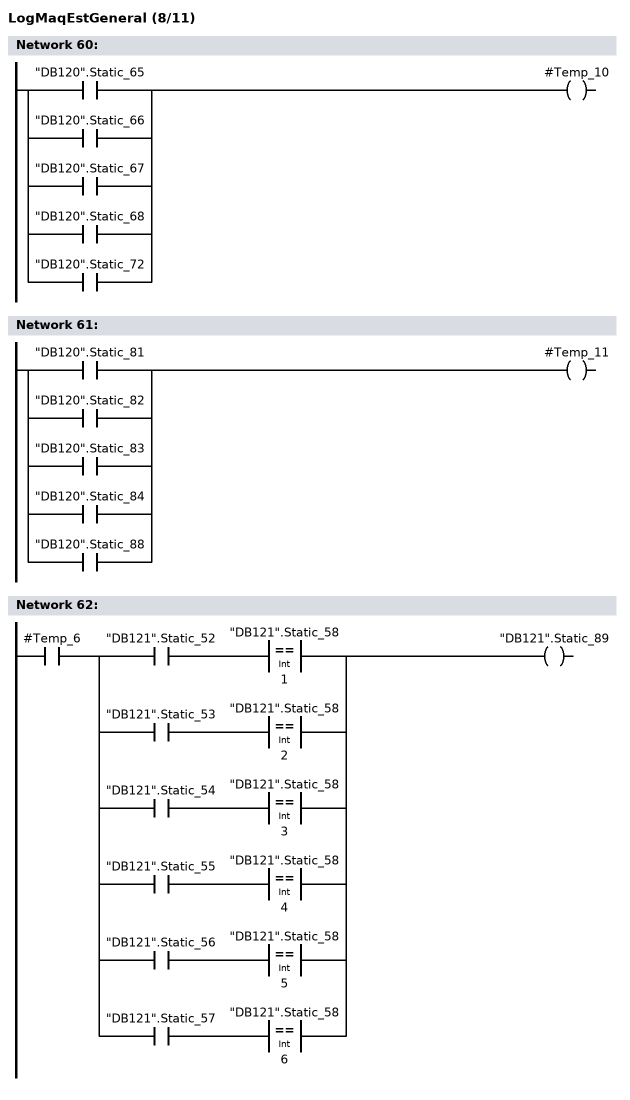
   RUNG wire#powerrail
      Contact( "DB120".Static_65 )
      wire#w1
      Coil( #Temp_10 )
   END_RUNG
   RUNG wire#powerrail
      Contact( "DB120".Static_66 )
   END_RUNG wire#w1
   RUNG wire#powerrail
      Contact( "DB120".Static_67 )
   END_RUNG wire#w1
   RUNG wire#powerrail
      Contact( "DB120".Static_68 )
   END_RUNG wire#w1
   RUNG wire#powerrail
      Contact( "DB120".Static_72 )
   END_RUNG wire#w1
   // the same network as SCL:
   #Temp_10 := "DB120".Static_65 OR "DB120".Static_66 OR "DB120".Static_67 OR "DB120".Static_68 OR "DB120".Static_72;
END_REGION

REGION Network 61
   RUNG wire#powerrail
      Contact( "DB120".Static_81 )
      wire#w1
      Coil( #Temp_11 )
   END_RUNG
   RUNG wire#powerrail
      Contact( "DB120".Static_82 )
   END_RUNG wire#w1
   RUNG wire#powerrail
      Contact( "DB120".Static_83 )
   END_RUNG wire#w1
   RUNG wire#powerrail
      Contact( "DB120".Static_84 )
   END_RUNG wire#w1
   RUNG wire#powerrail
      Contact( "DB120".Static_88 )
   END_RUNG wire#w1
   // the same network as SCL:
   #Temp_11 := "DB120".Static_81 OR "DB120".Static_82 OR "DB120".Static_83 OR "DB120".Static_84 OR "DB120".Static_88;
END_REGION

REGION Network 62
   "DB121".Static_89 := #Temp_6 AND (("DB121".Static_52 AND ("DB121".Static_58 = 1)) OR ("DB121".Static_53 AND ("DB121".Static_58 = 2)) OR ("DB121".Static_54 AND ("DB121".Static_58 = 3)) OR ("DB121".Static_55 AND ("DB121".Static_58 = 4)) OR ("DB121".Static_56 AND ("DB121".Static_58 = 5)) OR ("DB121".Static_57 AND ("DB121".Static_58 = 6)));
END_REGION

REGION Network 63
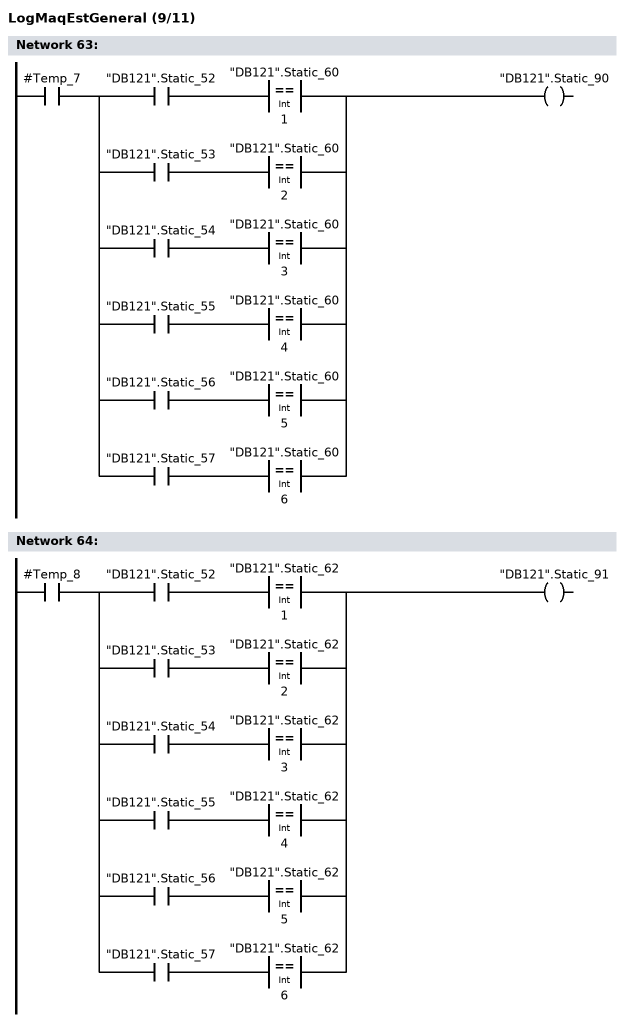
   "DB121".Static_90 := #Temp_7 AND (("DB121".Static_52 AND ("DB121".Static_60 = 1)) OR ("DB121".Static_53 AND ("DB121".Static_60 = 2)) OR ("DB121".Static_54 AND ("DB121".Static_60 = 3)) OR ("DB121".Static_55 AND ("DB121".Static_60 = 4)) OR ("DB121".Static_56 AND ("DB121".Static_60 = 5)) OR ("DB121".Static_57 AND ("DB121".Static_60 = 6)));
END_REGION

REGION Network 64
   "DB121".Static_91 := #Temp_8 AND (("DB121".Static_52 AND ("DB121".Static_62 = 1)) OR ("DB121".Static_53 AND ("DB121".Static_62 = 2)) OR ("DB121".Static_54 AND ("DB121".Static_62 = 3)) OR ("DB121".Static_55 AND ("DB121".Static_62 = 4)) OR ("DB121".Static_56 AND ("DB121".Static_62 = 5)) OR ("DB121".Static_57 AND ("DB121".Static_62 = 6)));
END_REGION

REGION Network 65
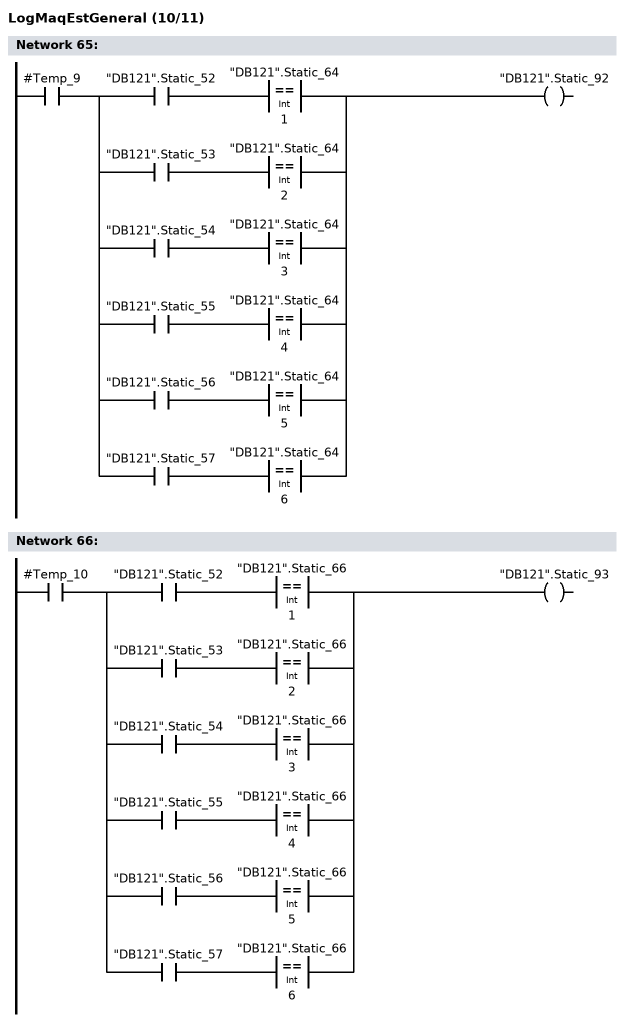
   "DB121".Static_92 := #Temp_9 AND (("DB121".Static_52 AND ("DB121".Static_64 = 1)) OR ("DB121".Static_53 AND ("DB121".Static_64 = 2)) OR ("DB121".Static_54 AND ("DB121".Static_64 = 3)) OR ("DB121".Static_55 AND ("DB121".Static_64 = 4)) OR ("DB121".Static_56 AND ("DB121".Static_64 = 5)) OR ("DB121".Static_57 AND ("DB121".Static_64 = 6)));
END_REGION

REGION Network 66
   "DB121".Static_93 := #Temp_10 AND (("DB121".Static_52 AND ("DB121".Static_66 = 1)) OR ("DB121".Static_53 AND ("DB121".Static_66 = 2)) OR ("DB121".Static_54 AND ("DB121".Static_66 = 3)) OR ("DB121".Static_55 AND ("DB121".Static_66 = 4)) OR ("DB121".Static_56 AND ("DB121".Static_66 = 5)) OR ("DB121".Static_57 AND ("DB121".Static_66 = 6)));
END_REGION

REGION Network 67
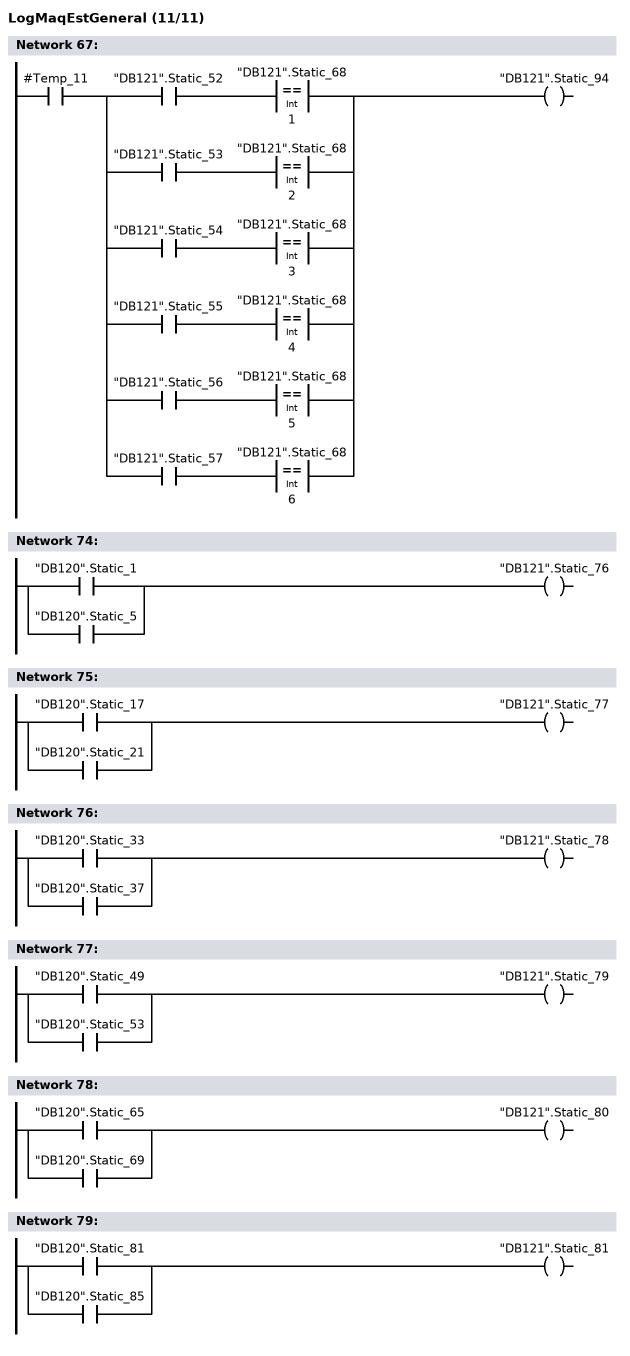
   "DB121".Static_94 := #Temp_11 AND (("DB121".Static_52 AND ("DB121".Static_68 = 1)) OR ("DB121".Static_53 AND ("DB121".Static_68 = 2)) OR ("DB121".Static_54 AND ("DB121".Static_68 = 3)) OR ("DB121".Static_55 AND ("DB121".Static_68 = 4)) OR ("DB121".Static_56 AND ("DB121".Static_68 = 5)) OR ("DB121".Static_57 AND ("DB121".Static_68 = 6)));
END_REGION

REGION Network 68 (STL)
         A(;
         L     "DB125".Static_1;
         L     1;
         ==R;
         );
         AN    "DB88".Static_12;
         O;
         A(;
         L     "DB125".Static_2;
         L     1;
         ==R;
         );
         AN    "DB88".Static_13;
         O;
         A(;
         L     "DB125".Static_3;
         L     1;
         ==R;
         );
         AN    "DB88".Static_14;
         O;
         A(;
         L     "DB125".Static_4;
         L     1;
         ==R;
         );
         AN    "DB88".Static_15;
         O;
         A(;
         L     "DB125".Static_5;
         L     1;
         ==R;
         );
         AN    "DB88".Static_16;
         O;
         A(;
         L     "DB125".Static_6;
         L     1;
         ==R;
         );
         AN    "DB88".Static_17;
         =     "DB121".Static_82;
END_REGION

REGION Network 69 (STL)
         A(;
         L     "DB125".Static_1;
         L     2;
         ==R;
         );
         AN    "DB88".Static_12;
         O;
         A(;
         L     "DB125".Static_2;
         L     2;
         ==R;
         );
         AN    "DB88".Static_13;
         O;
         A(;
         L     "DB125".Static_3;
         L     2;
         ==R;
         );
         AN    "DB88".Static_14;
         O;
         A(;
         L     "DB125".Static_4;
         L     2;
         ==R;
         );
         AN    "DB88".Static_15;
         O;
         A(;
         L     "DB125".Static_5;
         L     2;
         ==R;
         );
         AN    "DB88".Static_16;
         A(;
         L     "DB125".Static_6;
         L     2;
         ==R;
         );
         AN    "DB88".Static_17;
         =     "DB121".Static_83;
END_REGION

REGION Network 70 (STL)
         A(;
         L     "DB125".Static_1;
         L     3;
         ==R;
         );
         AN    "DB88".Static_12;
         O;
         A(;
         L     "DB125".Static_2;
         L     3;
         ==R;
         );
         AN    "DB88".Static_13;
         O;
         A(;
         L     "DB125".Static_3;
         L     3;
         ==R;
         );
         AN    "DB88".Static_14;
         O;
         A(;
         L     "DB125".Static_4;
         L     3;
         ==R;
         );
         AN    "DB88".Static_15;
         O;
         A(;
         L     "DB125".Static_5;
         L     3;
         ==R;
         );
         AN    "DB88".Static_16;
         O;
         A(;
         L     "DB125".Static_6;
         L     3;
         ==R;
         );
         AN    "DB88".Static_17;
         =     "DB121".Static_84;
END_REGION

REGION Network 71 (STL)
         A(;
         L     "DB125".Static_1;
         L     4;
         ==R;
         );
         AN    "DB88".Static_12;
         O;
         A(;
         L     "DB125".Static_2;
         L     4;
         ==R;
         );
         AN    "DB88".Static_13;
         O;
         A(;
         L     "DB125".Static_3;
         L     4;
         ==R;
         );
         AN    "DB88".Static_14;
         O;
         A(;
         L     "DB125".Static_4;
         L     4;
         ==R;
         );
         AN    "DB88".Static_15;
         O;
         A(;
         L     "DB125".Static_5;
         L     4;
         ==R;
         );
         AN    "DB88".Static_16;
         O;
         A(;
         L     "DB125".Static_6;
         L     4;
         ==R;
         );
         AN    "DB88".Static_17;
         =     "DB121".Static_85;
END_REGION

REGION Network 72 (STL)
         A(;
         L     "DB125".Static_1;
         L     5;
         ==R;
         );
         AN    "DB88".Static_12;
         O;
         A(;
         L     "DB125".Static_2;
         L     5;
         ==R;
         );
         AN    "DB88".Static_13;
         O;
         A(;
         L     "DB125".Static_3;
         L     5;
         ==R;
         );
         AN    "DB88".Static_14;
         O;
         A(;
         L     "DB125".Static_4;
         L     5;
         ==R;
         );
         AN    "DB88".Static_15;
         O;
         A(;
         L     "DB125".Static_5;
         L     5;
         ==R;
         );
         AN    "DB88".Static_16;
         O;
         A(;
         L     "DB125".Static_6;
         L     5;
         ==R;
         );
         AN    "DB88".Static_17;
         =     "DB121".Static_86;
END_REGION

REGION Network 73 (STL)
         A(;
         L     "DB125".Static_1;
         L     6;
         ==R;
         );
         AN    "DB88".Static_12;
         O;
         A(;
         L     "DB125".Static_2;
         L     6;
         ==R;
         );
         AN    "DB88".Static_13;
         O;
         A(;
         L     "DB125".Static_3;
         L     6;
         ==R;
         );
         AN    "DB88".Static_14;
         O;
         A(;
         L     "DB125".Static_4;
         L     6;
         ==R;
         );
         AN    "DB88".Static_15;
         O;
         A(;
         L     "DB125".Static_5;
         L     6;
         ==R;
         );
         AN    "DB88".Static_16;
         O;
         A(;
         L     "DB125".Static_6;
         L     6;
         ==R;
         );
         AN    "DB88".Static_17;
         =     "DB121".Static_87;
END_REGION

REGION Network 74
   RUNG wire#powerrail
      Contact( "DB120".Static_1 )
      wire#w1
      Coil( "DB121".Static_76 )
   END_RUNG
   RUNG wire#powerrail
      Contact( "DB120".Static_5 )
   END_RUNG wire#w1
   // the same network as SCL:
   "DB121".Static_76 := "DB120".Static_1 OR "DB120".Static_5;
END_REGION

REGION Network 75
   RUNG wire#powerrail
      Contact( "DB120".Static_17 )
      wire#w1
      Coil( "DB121".Static_77 )
   END_RUNG
   RUNG wire#powerrail
      Contact( "DB120".Static_21 )
   END_RUNG wire#w1
   // the same network as SCL:
   "DB121".Static_77 := "DB120".Static_17 OR "DB120".Static_21;
END_REGION

REGION Network 76
   RUNG wire#powerrail
      Contact( "DB120".Static_33 )
      wire#w1
      Coil( "DB121".Static_78 )
   END_RUNG
   RUNG wire#powerrail
      Contact( "DB120".Static_37 )
   END_RUNG wire#w1
   // the same network as SCL:
   "DB121".Static_78 := "DB120".Static_33 OR "DB120".Static_37;
END_REGION

REGION Network 77
   RUNG wire#powerrail
      Contact( "DB120".Static_49 )
      wire#w1
      Coil( "DB121".Static_79 )
   END_RUNG
   RUNG wire#powerrail
      Contact( "DB120".Static_53 )
   END_RUNG wire#w1
   // the same network as SCL:
   "DB121".Static_79 := "DB120".Static_49 OR "DB120".Static_53;
END_REGION

REGION Network 78
   RUNG wire#powerrail
      Contact( "DB120".Static_65 )
      wire#w1
      Coil( "DB121".Static_80 )
   END_RUNG
   RUNG wire#powerrail
      Contact( "DB120".Static_69 )
   END_RUNG wire#w1
   // the same network as SCL:
   "DB121".Static_80 := "DB120".Static_65 OR "DB120".Static_69;
END_REGION

REGION Network 79
   RUNG wire#powerrail
      Contact( "DB120".Static_81 )
      wire#w1
      Coil( "DB121".Static_81 )
   END_RUNG
   RUNG wire#powerrail
      Contact( "DB120".Static_85 )
   END_RUNG wire#w1
   // the same network as SCL:
   "DB121".Static_81 := "DB120".Static_81 OR "DB120".Static_85;
END_REGION
END_FUNCTION

FUNCTION "CalcEst1" : Void   // FC36, LAD
{ S7_Optimized_Access := 'FALSE' }
VERSION : 0.1
   VAR_TEMP   // added for the SCL form of the ladder/FBD networks
      _w1 : Bool;
   END_VAR
BEGIN

REGION Network 1
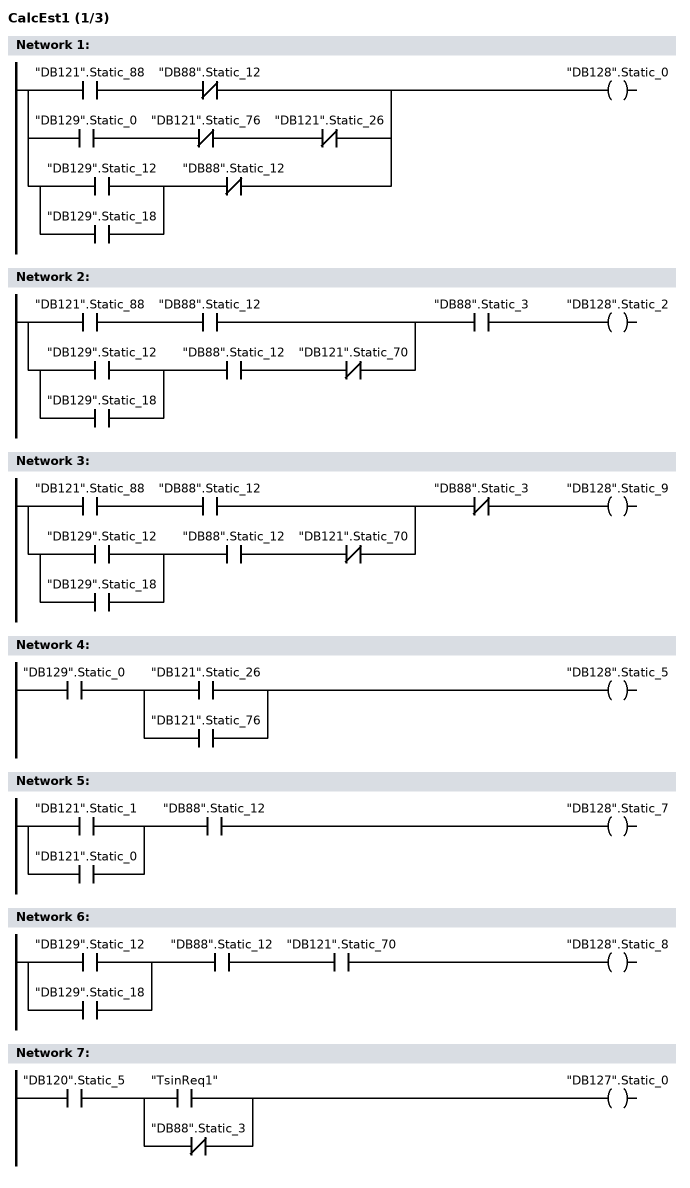
   RUNG wire#powerrail
      Contact( "DB121".Static_88 )
      I_Contact( "DB88".Static_12 )
      wire#w1
      Coil( "DB128".Static_0 )
   END_RUNG
   RUNG wire#powerrail
      Contact( "DB129".Static_0 )
      I_Contact( "DB121".Static_76 )
      I_Contact( "DB121".Static_26 )
   END_RUNG wire#w1
   RUNG wire#powerrail
      Contact( "DB129".Static_12 )
      wire#w2
      I_Contact( "DB88".Static_12 )
   END_RUNG wire#w1
   RUNG wire#powerrail
      Contact( "DB129".Static_18 )
   END_RUNG wire#w2
   // the same network as SCL:
   "DB128".Static_0 := ("DB121".Static_88 AND NOT "DB88".Static_12) OR ("DB129".Static_0 AND NOT "DB121".Static_76 AND NOT "DB121".Static_26) OR (("DB129".Static_12 OR "DB129".Static_18) AND NOT "DB88".Static_12);
END_REGION

REGION Network 2
   RUNG wire#powerrail
      Contact( "DB121".Static_88 )
      Contact( "DB88".Static_12 )
      wire#w1
      Contact( "DB88".Static_3 )
      Coil( "DB128".Static_2 )
   END_RUNG
   RUNG wire#powerrail
      Contact( "DB129".Static_12 )
      wire#w2
      Contact( "DB88".Static_12 )
      I_Contact( "DB121".Static_70 )
   END_RUNG wire#w1
   RUNG wire#powerrail
      Contact( "DB129".Static_18 )
   END_RUNG wire#w2
   // the same network as SCL:
   "DB128".Static_2 := (("DB121".Static_88 AND "DB88".Static_12) OR (("DB129".Static_12 OR "DB129".Static_18) AND "DB88".Static_12 AND NOT "DB121".Static_70)) AND "DB88".Static_3;
END_REGION

REGION Network 3
   RUNG wire#powerrail
      Contact( "DB121".Static_88 )
      Contact( "DB88".Static_12 )
      wire#w1
      I_Contact( "DB88".Static_3 )
      Coil( "DB128".Static_9 )
   END_RUNG
   RUNG wire#powerrail
      Contact( "DB129".Static_12 )
      wire#w2
      Contact( "DB88".Static_12 )
      I_Contact( "DB121".Static_70 )
   END_RUNG wire#w1
   RUNG wire#powerrail
      Contact( "DB129".Static_18 )
   END_RUNG wire#w2
   // the same network as SCL:
   "DB128".Static_9 := (("DB121".Static_88 AND "DB88".Static_12) OR (("DB129".Static_12 OR "DB129".Static_18) AND "DB88".Static_12 AND NOT "DB121".Static_70)) AND NOT "DB88".Static_3;
END_REGION

REGION Network 4
   "DB128".Static_5 := "DB129".Static_0 AND ("DB121".Static_26 OR "DB121".Static_76);
END_REGION

REGION Network 5
   RUNG wire#powerrail
      Contact( "DB121".Static_1 )
      wire#w1
      Contact( "DB88".Static_12 )
      Coil( "DB128".Static_7 )
   END_RUNG
   RUNG wire#powerrail
      Contact( "DB121".Static_0 )
   END_RUNG wire#w1
   // the same network as SCL:
   "DB128".Static_7 := ("DB121".Static_1 OR "DB121".Static_0) AND "DB88".Static_12;
END_REGION

REGION Network 6
   RUNG wire#powerrail
      Contact( "DB129".Static_12 )
      wire#w1
      Contact( "DB88".Static_12 )
      Contact( "DB121".Static_70 )
      Coil( "DB128".Static_8 )
   END_RUNG
   RUNG wire#powerrail
      Contact( "DB129".Static_18 )
   END_RUNG wire#w1
   // the same network as SCL:
   "DB128".Static_8 := ("DB129".Static_12 OR "DB129".Static_18) AND "DB88".Static_12 AND "DB121".Static_70;
END_REGION

REGION Network 7
   "DB127".Static_0 := "DB120".Static_5 AND ("TsinReq1" OR NOT "DB88".Static_3);
END_REGION

REGION Network 8
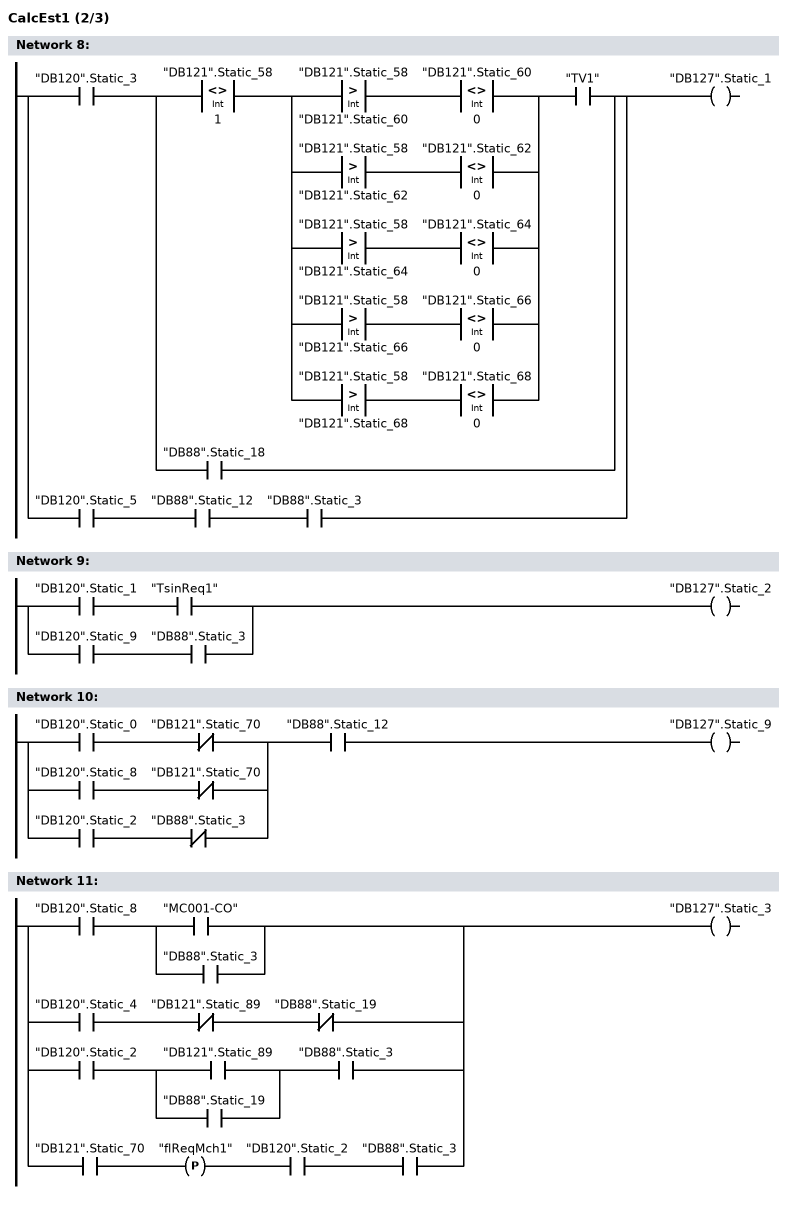
   "DB127".Static_1 := ("DB120".Static_3 AND ((("DB121".Static_58 <> 1) AND ((("DB121".Static_58 > "DB121".Static_60) AND ("DB121".Static_60 <> 0)) OR (("DB121".Static_58 > "DB121".Static_62) AND ("DB121".Static_62 <> 0)) OR (("DB121".Static_58 > "DB121".Static_64) AND ("DB121".Static_64 <> 0)) OR (("DB121".Static_58 > "DB121".Static_66) AND ("DB121".Static_66 <> 0)) OR (("DB121".Static_58 > "DB121".Static_68) AND ("DB121".Static_68 <> 0))) AND "TV1") OR "DB88".Static_18)) OR ("DB120".Static_5 AND "DB88".Static_12 AND "DB88".Static_3);
END_REGION

REGION Network 9
   RUNG wire#powerrail
      Contact( "DB120".Static_1 )
      Contact( "TsinReq1" )
      wire#w1
      Coil( "DB127".Static_2 )
   END_RUNG
   RUNG wire#powerrail
      Contact( "DB120".Static_9 )
      Contact( "DB88".Static_3 )
   END_RUNG wire#w1
   // the same network as SCL:
   "DB127".Static_2 := ("DB120".Static_1 AND "TsinReq1") OR ("DB120".Static_9 AND "DB88".Static_3);
END_REGION

REGION Network 10
   RUNG wire#powerrail
      Contact( "DB120".Static_0 )
      I_Contact( "DB121".Static_70 )
      wire#w1
      Contact( "DB88".Static_12 )
      Coil( "DB127".Static_9 )
   END_RUNG
   RUNG wire#powerrail
      Contact( "DB120".Static_8 )
      I_Contact( "DB121".Static_70 )
   END_RUNG wire#w1
   RUNG wire#powerrail
      Contact( "DB120".Static_2 )
      I_Contact( "DB88".Static_3 )
   END_RUNG wire#w1
   // the same network as SCL:
   "DB127".Static_9 := (("DB120".Static_0 AND NOT "DB121".Static_70) OR ("DB120".Static_8 AND NOT "DB121".Static_70) OR ("DB120".Static_2 AND NOT "DB88".Static_3)) AND "DB88".Static_12;
END_REGION

REGION Network 11
   #_w1 := "DB121".Static_70 AND NOT "flReqMch1";   // rising edge
   "flReqMch1" := "DB121".Static_70;
   "DB127".Static_3 := ("DB120".Static_8 AND ("MC001-CO" OR "DB88".Static_3)) OR ("DB120".Static_4 AND NOT "DB121".Static_89 AND NOT "DB88".Static_19) OR ("DB120".Static_2 AND ("DB121".Static_89 OR "DB88".Static_19) AND "DB88".Static_3) OR (#_w1 AND "DB120".Static_2 AND "DB88".Static_3);
END_REGION

REGION Network 12
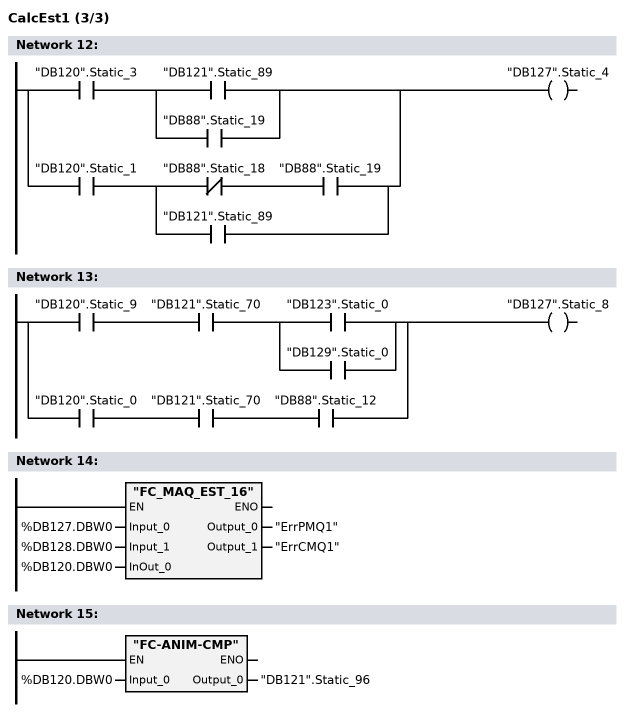
   "DB127".Static_4 := ("DB120".Static_3 AND ("DB121".Static_89 OR "DB88".Static_19)) OR ("DB120".Static_1 AND ("DB121".Static_89 OR (NOT "DB88".Static_18 AND "DB88".Static_19)));
END_REGION

REGION Network 13
   "DB127".Static_8 := ("DB120".Static_9 AND "DB121".Static_70 AND ("DB123".Static_0 OR "DB129".Static_0)) OR ("DB120".Static_0 AND "DB121".Static_70 AND "DB88".Static_12);
END_REGION

REGION Network 14
   RUNG wire#powerrail
      "FC_MAQ_EST_16"(Input_0 := %DB127.DBW0, Input_1 := %DB128.DBW0, Output_0 => "ErrPMQ1", Output_1 => "ErrCMQ1", InOut_0 := %DB120.DBW0)
   END_RUNG
   // the same network as SCL:
   "FC_MAQ_EST_16"(Input_0 := %DB127.DBW0,
                   Input_1 := %DB128.DBW0,
                   InOut_0 := %DB120.DBW0,
                   Output_0 => "ErrPMQ1",
                   Output_1 => "ErrCMQ1");
END_REGION

REGION Network 15
   RUNG wire#powerrail
      "FC-ANIM-CMP"(Input_0 := %DB120.DBW0, Output_0 => "DB121".Static_96)
   END_RUNG
   // the same network as SCL:
   "FC-ANIM-CMP"(Input_0 := %DB120.DBW0, Output_0 => "DB121".Static_96);
END_REGION
END_FUNCTION

FUNCTION "CalcEst2" : Void   // FC37, LAD
{ S7_Optimized_Access := 'FALSE' }
VERSION : 0.1
   VAR_TEMP   // added for the SCL form of the ladder/FBD networks
      _w1 : Bool;
   END_VAR
BEGIN

REGION Network 1
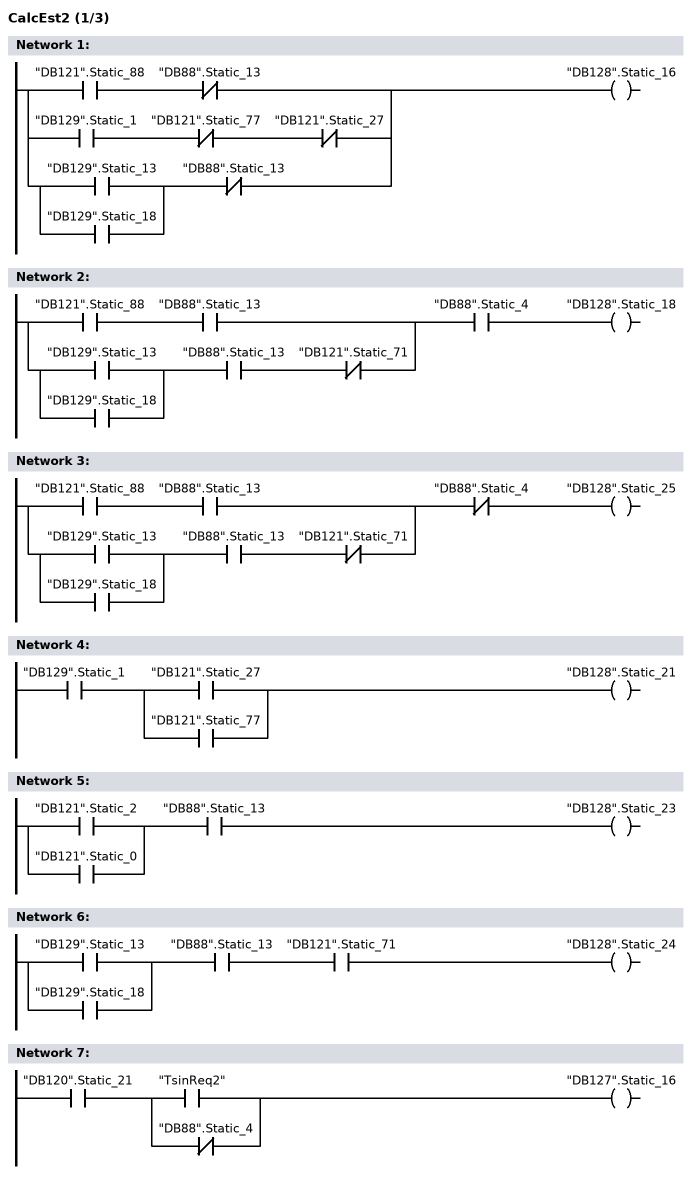
   RUNG wire#powerrail
      Contact( "DB121".Static_88 )
      I_Contact( "DB88".Static_13 )
      wire#w1
      Coil( "DB128".Static_16 )
   END_RUNG
   RUNG wire#powerrail
      Contact( "DB129".Static_1 )
      I_Contact( "DB121".Static_77 )
      I_Contact( "DB121".Static_27 )
   END_RUNG wire#w1
   RUNG wire#powerrail
      Contact( "DB129".Static_13 )
      wire#w2
      I_Contact( "DB88".Static_13 )
   END_RUNG wire#w1
   RUNG wire#powerrail
      Contact( "DB129".Static_18 )
   END_RUNG wire#w2
   // the same network as SCL:
   "DB128".Static_16 := ("DB121".Static_88 AND NOT "DB88".Static_13) OR ("DB129".Static_1 AND NOT "DB121".Static_77 AND NOT "DB121".Static_27) OR (("DB129".Static_13 OR "DB129".Static_18) AND NOT "DB88".Static_13);
END_REGION

REGION Network 2
   RUNG wire#powerrail
      Contact( "DB121".Static_88 )
      Contact( "DB88".Static_13 )
      wire#w1
      Contact( "DB88".Static_4 )
      Coil( "DB128".Static_18 )
   END_RUNG
   RUNG wire#powerrail
      Contact( "DB129".Static_13 )
      wire#w2
      Contact( "DB88".Static_13 )
      I_Contact( "DB121".Static_71 )
   END_RUNG wire#w1
   RUNG wire#powerrail
      Contact( "DB129".Static_18 )
   END_RUNG wire#w2
   // the same network as SCL:
   "DB128".Static_18 := (("DB121".Static_88 AND "DB88".Static_13) OR (("DB129".Static_13 OR "DB129".Static_18) AND "DB88".Static_13 AND NOT "DB121".Static_71)) AND "DB88".Static_4;
END_REGION

REGION Network 3
   RUNG wire#powerrail
      Contact( "DB121".Static_88 )
      Contact( "DB88".Static_13 )
      wire#w1
      I_Contact( "DB88".Static_4 )
      Coil( "DB128".Static_25 )
   END_RUNG
   RUNG wire#powerrail
      Contact( "DB129".Static_13 )
      wire#w2
      Contact( "DB88".Static_13 )
      I_Contact( "DB121".Static_71 )
   END_RUNG wire#w1
   RUNG wire#powerrail
      Contact( "DB129".Static_18 )
   END_RUNG wire#w2
   // the same network as SCL:
   "DB128".Static_25 := (("DB121".Static_88 AND "DB88".Static_13) OR (("DB129".Static_13 OR "DB129".Static_18) AND "DB88".Static_13 AND NOT "DB121".Static_71)) AND NOT "DB88".Static_4;
END_REGION

REGION Network 4
   "DB128".Static_21 := "DB129".Static_1 AND ("DB121".Static_27 OR "DB121".Static_77);
END_REGION

REGION Network 5
   RUNG wire#powerrail
      Contact( "DB121".Static_2 )
      wire#w1
      Contact( "DB88".Static_13 )
      Coil( "DB128".Static_23 )
   END_RUNG
   RUNG wire#powerrail
      Contact( "DB121".Static_0 )
   END_RUNG wire#w1
   // the same network as SCL:
   "DB128".Static_23 := ("DB121".Static_2 OR "DB121".Static_0) AND "DB88".Static_13;
END_REGION

REGION Network 6
   RUNG wire#powerrail
      Contact( "DB129".Static_13 )
      wire#w1
      Contact( "DB88".Static_13 )
      Contact( "DB121".Static_71 )
      Coil( "DB128".Static_24 )
   END_RUNG
   RUNG wire#powerrail
      Contact( "DB129".Static_18 )
   END_RUNG wire#w1
   // the same network as SCL:
   "DB128".Static_24 := ("DB129".Static_13 OR "DB129".Static_18) AND "DB88".Static_13 AND "DB121".Static_71;
END_REGION

REGION Network 7
   "DB127".Static_16 := "DB120".Static_21 AND ("TsinReq2" OR NOT "DB88".Static_4);
END_REGION

REGION Network 8
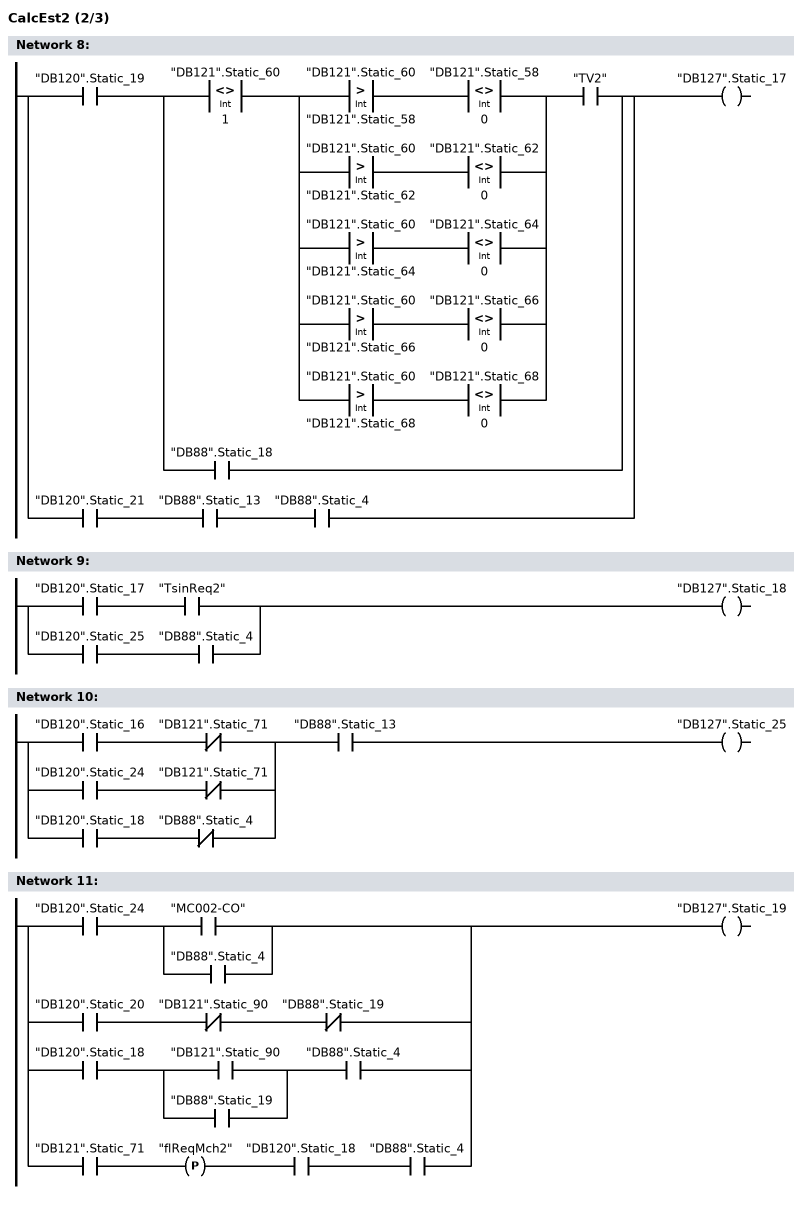
   "DB127".Static_17 := ("DB120".Static_19 AND ((("DB121".Static_60 <> 1) AND ((("DB121".Static_60 > "DB121".Static_58) AND ("DB121".Static_58 <> 0)) OR (("DB121".Static_60 > "DB121".Static_62) AND ("DB121".Static_62 <> 0)) OR (("DB121".Static_60 > "DB121".Static_64) AND ("DB121".Static_64 <> 0)) OR (("DB121".Static_60 > "DB121".Static_66) AND ("DB121".Static_66 <> 0)) OR (("DB121".Static_60 > "DB121".Static_68) AND ("DB121".Static_68 <> 0))) AND "TV2") OR "DB88".Static_18)) OR ("DB120".Static_21 AND "DB88".Static_13 AND "DB88".Static_4);
END_REGION

REGION Network 9
   RUNG wire#powerrail
      Contact( "DB120".Static_17 )
      Contact( "TsinReq2" )
      wire#w1
      Coil( "DB127".Static_18 )
   END_RUNG
   RUNG wire#powerrail
      Contact( "DB120".Static_25 )
      Contact( "DB88".Static_4 )
   END_RUNG wire#w1
   // the same network as SCL:
   "DB127".Static_18 := ("DB120".Static_17 AND "TsinReq2") OR ("DB120".Static_25 AND "DB88".Static_4);
END_REGION

REGION Network 10
   RUNG wire#powerrail
      Contact( "DB120".Static_16 )
      I_Contact( "DB121".Static_71 )
      wire#w1
      Contact( "DB88".Static_13 )
      Coil( "DB127".Static_25 )
   END_RUNG
   RUNG wire#powerrail
      Contact( "DB120".Static_24 )
      I_Contact( "DB121".Static_71 )
   END_RUNG wire#w1
   RUNG wire#powerrail
      Contact( "DB120".Static_18 )
      I_Contact( "DB88".Static_4 )
   END_RUNG wire#w1
   // the same network as SCL:
   "DB127".Static_25 := (("DB120".Static_16 AND NOT "DB121".Static_71) OR ("DB120".Static_24 AND NOT "DB121".Static_71) OR ("DB120".Static_18 AND NOT "DB88".Static_4)) AND "DB88".Static_13;
END_REGION

REGION Network 11
   #_w1 := "DB121".Static_71 AND NOT "flReqMch2";   // rising edge
   "flReqMch2" := "DB121".Static_71;
   "DB127".Static_19 := ("DB120".Static_24 AND ("MC002-CO" OR "DB88".Static_4)) OR ("DB120".Static_20 AND NOT "DB121".Static_90 AND NOT "DB88".Static_19) OR ("DB120".Static_18 AND ("DB121".Static_90 OR "DB88".Static_19) AND "DB88".Static_4) OR (#_w1 AND "DB120".Static_18 AND "DB88".Static_4);
END_REGION

REGION Network 12
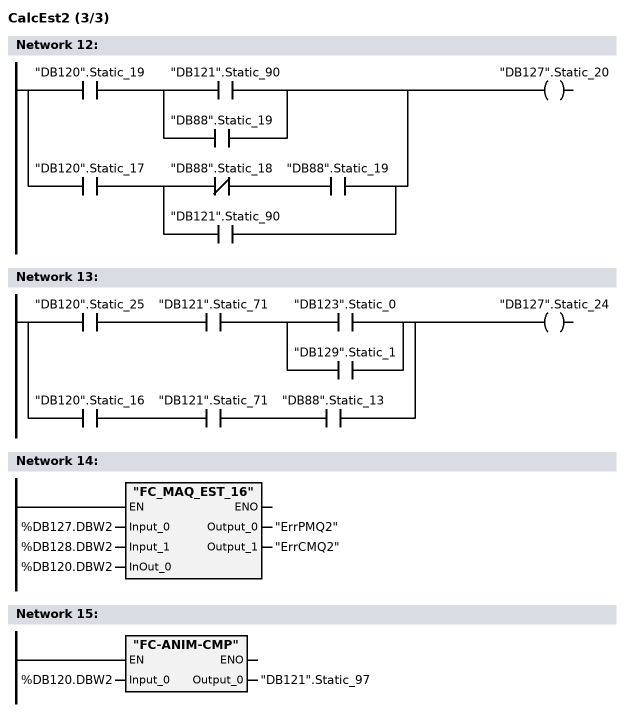
   "DB127".Static_20 := ("DB120".Static_19 AND ("DB121".Static_90 OR "DB88".Static_19)) OR ("DB120".Static_17 AND ("DB121".Static_90 OR (NOT "DB88".Static_18 AND "DB88".Static_19)));
END_REGION

REGION Network 13
   "DB127".Static_24 := ("DB120".Static_25 AND "DB121".Static_71 AND ("DB123".Static_0 OR "DB129".Static_1)) OR ("DB120".Static_16 AND "DB121".Static_71 AND "DB88".Static_13);
END_REGION

REGION Network 14
   RUNG wire#powerrail
      "FC_MAQ_EST_16"(Input_0 := %DB127.DBW2, Input_1 := %DB128.DBW2, Output_0 => "ErrPMQ2", Output_1 => "ErrCMQ2", InOut_0 := %DB120.DBW2)
   END_RUNG
   // the same network as SCL:
   "FC_MAQ_EST_16"(Input_0 := %DB127.DBW2,
                   Input_1 := %DB128.DBW2,
                   InOut_0 := %DB120.DBW2,
                   Output_0 => "ErrPMQ2",
                   Output_1 => "ErrCMQ2");
END_REGION

REGION Network 15
   RUNG wire#powerrail
      "FC-ANIM-CMP"(Input_0 := %DB120.DBW2, Output_0 => "DB121".Static_97)
   END_RUNG
   // the same network as SCL:
   "FC-ANIM-CMP"(Input_0 := %DB120.DBW2, Output_0 => "DB121".Static_97);
END_REGION
END_FUNCTION

FUNCTION "CalcEst3" : Void   // FC38, LAD
{ S7_Optimized_Access := 'FALSE' }
VERSION : 0.1
   VAR_TEMP   // added for the SCL form of the ladder/FBD networks
      _w1 : Bool;
   END_VAR
BEGIN

REGION Network 1
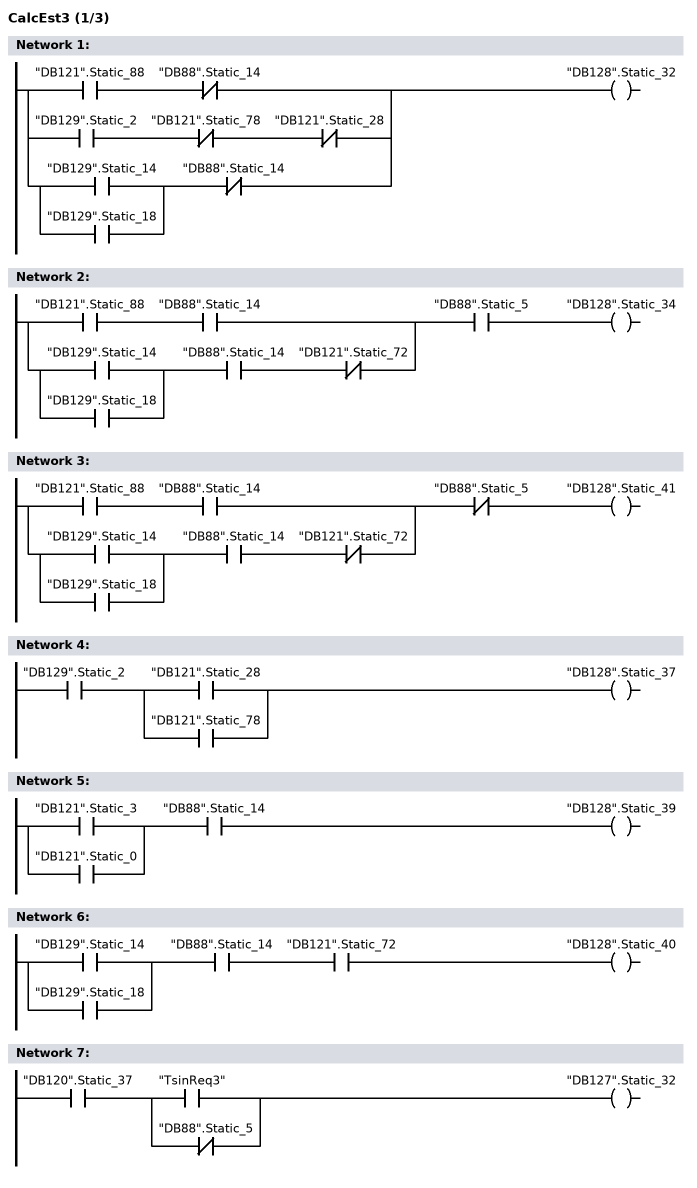
   RUNG wire#powerrail
      Contact( "DB121".Static_88 )
      I_Contact( "DB88".Static_14 )
      wire#w1
      Coil( "DB128".Static_32 )
   END_RUNG
   RUNG wire#powerrail
      Contact( "DB129".Static_2 )
      I_Contact( "DB121".Static_78 )
      I_Contact( "DB121".Static_28 )
   END_RUNG wire#w1
   RUNG wire#powerrail
      Contact( "DB129".Static_14 )
      wire#w2
      I_Contact( "DB88".Static_14 )
   END_RUNG wire#w1
   RUNG wire#powerrail
      Contact( "DB129".Static_18 )
   END_RUNG wire#w2
   // the same network as SCL:
   "DB128".Static_32 := ("DB121".Static_88 AND NOT "DB88".Static_14) OR ("DB129".Static_2 AND NOT "DB121".Static_78 AND NOT "DB121".Static_28) OR (("DB129".Static_14 OR "DB129".Static_18) AND NOT "DB88".Static_14);
END_REGION

REGION Network 2
   RUNG wire#powerrail
      Contact( "DB121".Static_88 )
      Contact( "DB88".Static_14 )
      wire#w1
      Contact( "DB88".Static_5 )
      Coil( "DB128".Static_34 )
   END_RUNG
   RUNG wire#powerrail
      Contact( "DB129".Static_14 )
      wire#w2
      Contact( "DB88".Static_14 )
      I_Contact( "DB121".Static_72 )
   END_RUNG wire#w1
   RUNG wire#powerrail
      Contact( "DB129".Static_18 )
   END_RUNG wire#w2
   // the same network as SCL:
   "DB128".Static_34 := (("DB121".Static_88 AND "DB88".Static_14) OR (("DB129".Static_14 OR "DB129".Static_18) AND "DB88".Static_14 AND NOT "DB121".Static_72)) AND "DB88".Static_5;
END_REGION

REGION Network 3
   RUNG wire#powerrail
      Contact( "DB121".Static_88 )
      Contact( "DB88".Static_14 )
      wire#w1
      I_Contact( "DB88".Static_5 )
      Coil( "DB128".Static_41 )
   END_RUNG
   RUNG wire#powerrail
      Contact( "DB129".Static_14 )
      wire#w2
      Contact( "DB88".Static_14 )
      I_Contact( "DB121".Static_72 )
   END_RUNG wire#w1
   RUNG wire#powerrail
      Contact( "DB129".Static_18 )
   END_RUNG wire#w2
   // the same network as SCL:
   "DB128".Static_41 := (("DB121".Static_88 AND "DB88".Static_14) OR (("DB129".Static_14 OR "DB129".Static_18) AND "DB88".Static_14 AND NOT "DB121".Static_72)) AND NOT "DB88".Static_5;
END_REGION

REGION Network 4
   "DB128".Static_37 := "DB129".Static_2 AND ("DB121".Static_28 OR "DB121".Static_78);
END_REGION

REGION Network 5
   RUNG wire#powerrail
      Contact( "DB121".Static_3 )
      wire#w1
      Contact( "DB88".Static_14 )
      Coil( "DB128".Static_39 )
   END_RUNG
   RUNG wire#powerrail
      Contact( "DB121".Static_0 )
   END_RUNG wire#w1
   // the same network as SCL:
   "DB128".Static_39 := ("DB121".Static_3 OR "DB121".Static_0) AND "DB88".Static_14;
END_REGION

REGION Network 6
   RUNG wire#powerrail
      Contact( "DB129".Static_14 )
      wire#w1
      Contact( "DB88".Static_14 )
      Contact( "DB121".Static_72 )
      Coil( "DB128".Static_40 )
   END_RUNG
   RUNG wire#powerrail
      Contact( "DB129".Static_18 )
   END_RUNG wire#w1
   // the same network as SCL:
   "DB128".Static_40 := ("DB129".Static_14 OR "DB129".Static_18) AND "DB88".Static_14 AND "DB121".Static_72;
END_REGION

REGION Network 7
   "DB127".Static_32 := "DB120".Static_37 AND ("TsinReq3" OR NOT "DB88".Static_5);
END_REGION

REGION Network 8